
         O(;
         L     #Temp_PV.PV_SetV.WarningUpperLimit;
         L     0.0;
         <=R;
         );
         O(;
         L     #Temp_PV.PV_SetV.Value;
         L     #Temp_PV.PV_SetV.WarningUpperLimit;
         +R;
         L     #Temp_PV.PV_ActV.Value;
         >R;
         );
         JC    gwon;

         L     4;
         T     #Temp_PV.PV_ActV.ValueState;

         JU    end;

   gwon: NOP   0;

   end:  NOP   0;
END_REGION

REGION Network 4: Detect fault levels
   ENDC: O(;
         L     #Temp_PV.PV_ActV.ValueState;
         L     1;
         AW;
         L     0;
         >I;
         );
         AN    #IO_Fault_Alarm_lowerL;
         S     #IO_Fault_Alarm_lowerL;
         S     #IO_New_Fault;

         O(;
         L     #Temp_PV.PV_ActV.ValueState;
         L     2;
         AW;
         L     0;
         >I;
         );
         AN    #IO_Fault_Warn_lowerL;
         S     #IO_Fault_Warn_lowerL;
         S     #IO_New_Fault;

         O(;
         L     #Temp_PV.PV_ActV.ValueState;
         L     4;
         AW;
         L     0;
         >I;
         );
         AN    #IO_Fault_Warn_upperL;
         S     #IO_Fault_Warn_upperL;
         S     #IO_New_Fault;

         O(;
         L     #Temp_PV.PV_ActV.ValueState;
         L     8;
         AW;
         L     0;
         >I;
         );
         AN    #IO_Fault_Alarm_upperL;
         S     #IO_Fault_Alarm_upperL;
         S     #IO_New_Fault;

         O     #IO_Fault_Alarm_lowerL;
         O     #IO_Fault_Alarm_upperL;
         S     #IO_Fault_Level_1;

         O     #IO_Fault_Warn_lowerL;
         O     #IO_Fault_Warn_upperL;
         S     #IO_Fault_Level_3;
END_REGION

REGION Network 5: Write actual value to DB
         CALL  BLKMOV
         ( SRCBLK  := #Temp_PV,
           RET_VAL := #RetVal,
           DSTBLK  := #Anyzeiger_PV
         );
END_REGION
END_FUNCTION

FUNCTION "FC920_PV_Calc_Act_Value" : Void   // FC920, STL
TITLE = Calculates the actual process value of a source
{ S7_Optimized_Access := 'FALSE' }
AUTHOR : HK
VERSION : 0.1
   VAR_INPUT
      IN_Act_Value_read : Bool;   // Read actual value 0 = NO, 1 = YES
      IN_Act_Value_ext : Bool;   // Get actual value from extern
      IN_Ext_Value : Real;   // External value DWord
      IN_Read_Double : Bool;   // Read double word value
      IN_FLT_Needful : Bool;   // Is a seperat fault identification needful?
      IN_FLT_Reset : Bool;
   END_VAR
   VAR_IN_OUT
      IO_Any_ArrayPV : ANY;
      IO_Fault_Sensor : Bool;
      IO_New_Fault : Bool;
      IO_FLT_Level_3 : Bool;
   END_VAR
   VAR_TEMP
      RetVal : Int;
      Anz_BytePV_Act : Int;
      DB_Nr_PV_Act : Int;
      Anyzeiger_Act : ANY;
      Anf_1_PV_Act : Byte;
      Anf_2_PV_Act : Word;
      Temp_PV : "UDT910_ProcessValue";
      Temp_ActV_Pointer : DWord;
      Temp_Fault_Sensor : Bool;
      Temp_CheckSensor : Bool;
   END_VAR
BEGIN

REGION Network 1: Read Array[No_Array] actual value conf. and actual value
         L;  // Pointer auf das Arrays
         LAR1;

         L     W[AR1, P#2.0];  // #Anz_Byte Baugruppe
         T     #Anz_BytePV_Act;

         L     W[AR1, P#4.0];
         T     #DB_Nr_PV_Act;  // DB no prozessvalue actual value

         L     B[AR1, P#7.0];
         T     #Anf_1_PV_Act;

         L     W[AR1, P#8.0];
         T     #Anf_2_PV_Act;  // Start DW prozessvalue actual value [0]

   //
         LAR1;
         L     16#1002;  // Bytes
         T     W[AR1, P#0.0];
         L     #Anz_BytePV_Act;  // Amount of bytes
         T     W[AR1, P#2.0];
         L     #DB_Nr_PV_Act;  // Block no,
         T     W[AR1, P#4.0];
         L     16#84;
         T     LB[AR1, P#6.0];
         L     #Anf_1_PV_Act;
         T     LB[AR1, P#7.0];
         L     #Anf_2_PV_Act;
         T     LW[AR1, P#8.0];

   //
         CALL  BLKMOV
         ( SRCBLK  := #Anyzeiger_Act,
           RET_VAL := #RetVal,
           DSTBLK  := #Temp_PV
         );
   //

   //------- Reset fault -----------------------
         A     #IN_FLT_Reset;
         ON    #IN_FLT_Needful;
         R     #IO_Fault_Sensor;
END_REGION

REGION Network 2: Reset process value
         L     0;
         T     #Temp_PV.PV_ActV.Value;
   //-----
         AN    #IN_Act_Value_read;
         JC    end6;
   //-------------------------------------------
         A     #IN_Act_Value_ext;  // Value is set external
         A     #IN_Act_Value_read;
         JC    extv;
   //-------------------------------------------
         L     #Temp_PV.PV_Conf_ActV.Address;
         L     0;
         ==I;
         JC    end6;
   //-----
END_REGION

REGION Network 3: Calculate actual value

         A     #IN_Act_Value_ext;  // Value is set external
         JC    extv;
   //-------------------------------------------

         L     #Temp_PV.PV_Conf_ActV.Address;
         SLD   3;
         T     #Temp_ActV_Pointer;

         AN    #IN_Read_Double;
         JC    word;
         L     PID[ #Temp_ActV_Pointer];
         T     #Temp_PV.PV_ActV.Value;
         JU    nw02;
   word: L     PIW[ #Temp_ActV_Pointer];
         ITD;
         DTR;
         T     #Temp_PV.PV_ActV.Value;
         JU    nw02;

   extv: L     #IN_Ext_Value;
         T     #Temp_PV.PV_ActV.Value;

   nw02: L     #Temp_PV.PV_Conf_ActV.Multiplier;
         L     0.0;
         ==R;
         JC    nw03;
         L     #Temp_PV.PV_ActV.Value;
         L     #Temp_PV.PV_Conf_ActV.OffsetSignal;
         ITD;
         DTR;
         -R;
         L     #Temp_PV.PV_Conf_ActV.Multiplier;
         /R;
         T     #Temp_PV.PV_ActV.Value;
END_REGION

REGION Network 4: Limit control sensor value if limits <> 0
   nw03: L     #Temp_PV.PV_Conf_ActV.MaxValueSensor;
         L     #Temp_PV.PV_Conf_ActV.MinValueSensor;
         OW;
         L     0;
         <>D;
         =     #Temp_CheckSensor;

         O(;
         L     #Temp_PV.PV_ActV.Value;
         L     #Temp_PV.PV_Conf_ActV.MaxValueSensor;
         >R;
         );
         O(;
         L     #Temp_PV.PV_ActV.Value;
         L     #Temp_PV.PV_Conf_ActV.MinValueSensor;
         <R;
         );
         A     #Temp_CheckSensor;
         =     #Temp_Fault_Sensor;

         AN    #IN_FLT_Needful;
         JC    ResetValue;

         A     #Temp_Fault_Sensor;
         AN    #IO_Fault_Sensor;
         S     #IO_Fault_Sensor;
         S     #IO_New_Fault;

         O     #IO_Fault_Sensor;
         A     #IN_FLT_Needful;
         S     #IO_FLT_Level_3;
         JU    ResetValue;

   NSepFault:NOP   0;
         A     #Temp_Fault_Sensor;
         =     #IO_Fault_Sensor;

   ResetValue:NOP   0;
         AN    #Temp_Fault_Sensor;
         JC    end6;
         L     0.0;
         T     #Temp_PV.PV_ActV.Value;
         JU    end6;
END_REGION

REGION Network 5: Write actual value to DB
   end6: CALL  BLKMOV
         ( SRCBLK  := #Temp_PV,
           RET_VAL := #RetVal,
           DSTBLK  := #Anyzeiger_Act
         );
END_REGION
END_FUNCTION

FUNCTION "CHCKPNCONN" : Void   // FC1001, SCL
{ S7_Optimized_Access := 'FALSE' }
VERSION : 0.1
   VAR_IN_OUT
      GOON : Bool;
      Active : Bool;
      Address : Hw_Io;
      PN_Request : Bool;
      PN_Fault : Bool;
      DONE : Bool;
   END_VAR
   VAR_TEMP
      SLZ_Header : Struct
         LENTHDR : Word;
         N_DR : Word;
      END_STRUCT;
      Dataset : "SZL-IDW#16#xy96_DataSet";
      ReturnValue : Word;
      ReturnValue_1 : Int;
      ReturnHW : Int;
      HW_Kennung : Hw_Io;
      TempAddress : Hw_Io;
      HW_KennungDevice : Hw_SubModule;
      variant_inout : Variant;
   END_VAR
BEGIN
   IF NOT #GOON THEN
       #DONE := false;
   END_IF;

   IF #Active THEN
       IF #GOON AND NOT #DONE THEN

           "PN_Get_DIAG".returnValue := GET_DIAG(MODE := "PN_Get_DIAG".diagMODE, LADDR := #Address,
                                                 CNT_DIAG => "PN_Get_DIAG".CountDiagDetails,
                                                 DIAG := "PN_Get_DIAG".Diag,
                                                 DETAIL :=#variant_inout);

           IF "Flag_Req_read_IO_Busy" = 0 THEN
               // Bearbeitung beendet
               #DONE := true;
               // Fehler wurde festgestellt
               IF ("PN_Get_DIAG".Diag.OwnState > 0)

               THEN
                   #PN_Fault := true;
                   #PN_Request := false;
               END_IF;
               // Fehler wurde behoben
               IF #PN_Fault AND ("PN_Get_DIAG".Diag.OwnState = 0)

               THEN
                   #PN_Request := true;//#PN_Fault;
                   #PN_Fault := false;
               END_IF;
           END_IF;
       END_IF;
   ELSE
       #DONE := #GOON;
   END_IF;
   // Zusätzlichen Ausgang schreiben
   // 
   #GOON := #DONE;



   // Unten ist der alte Code
   // IF #GoOn THEN
   //     #ReturnValue := INT_TO_WORD(RDSYSST(REQ := true, //"Flag_01_000_Hertz" ,
   //                                                                     SZL_ID := 16#0696,
   //                                                                     INDEX := DINT_TO_WORD(#Address),
   //                                                                     BUSY => "Flag_Req_read_DP1_Busy",
   //                                                                     SZL_HEADER => #SLZ_Header,
   //                                                                     DR => "PN_CON".Dataset));

   //     IF #ReturnValue <> 0 THEN
   //         IF (NOT "PN_CON".Dataset.IOStat.BaugruppeVorhanden) OR "PN_CON".Dataset.IOStat.BaugruppeDeaktiviert OR "PN_CON".Dataset.IOStat.BaugruppeNichtVerfuegbar THEN

   //             #PN_Fault := true;
   //             #PN_Request := false;
   //         END_IF;

   //         IF #PN_Fault AND "PN_CON".Dataset.IOStat.BaugruppeVorhanden AND NOT "PN_CON".Dataset.IOStat.BaugruppeDeaktiviert AND NOT "PN_CON".Dataset.IOStat.BaugruppeNichtVerfuegbar THEN
   //             #PN_Request := true;
   //             #PN_Fault := false;
   //         END_IF;
   //     END_IF;
   //     IF WORD_TO_INT(#ReturnValue) > 16#8000 THEN
   //             #PN_Fault := true;
   //     END_IF;
   // END_IF;
END_FUNCTION

FUNCTION "PNC_AI" : Void   // FC1002, SCL
{ S7_Optimized_Access := 'FALSE' }
VERSION : 0.1
   VAR_INPUT
      RequestAll : Bool;
      AcknowledgeFaults : Bool;
   END_VAR
   VAR_IN_OUT
      GOON : Bool;
   END_VAR
   VAR_TEMP
      t : Struct
         DONE : Bool;
         BUSY : Bool;
         ERROR : Bool;
         STATUS : DWord;
      END_STRUCT;
      MODULE : Int;
      ADDRESS : Word;
      MinIndex : Int;
      MaxIndex : Int;
      SLZ_Header : Struct
         LENTHDR : Word;
         N_DR : Word;
      END_STRUCT;
      Dataset : "SZL-IDW#16#xy96_DataSet";
      TempHWID : Hw_Io;
      ReturnValue : Int;
   END_VAR
   VAR CONSTANT
      IDM_Analogin_Default_Skalierung_Index : Int := 2;
      IDM_Analogin_Default_Skalierung_Length : Int := 4;
      IDM_Analogin_Default_Filterung_Index : Int := 3;
      IDM_Analogin_Default_Filterung_Length : Int := 2;
      IDM_Analogin_Default_Grenzen_Index : Int := 4;
      IDM_Analogin_Default_Grenzen_Length : Int := 12;
      IDM_Analogin_Default_8_X14_0_Index : Int := 1;
      IDM_Analogin_Default_8_X14_0_Length : Int := 64;
      IDM_Analogin_Temperature_Index : Int := 2;
      IDM_Analogin_Temperature_Length : Int := 5;
      IDM_Analogin_Temperature_8_Index : Int := 1;
      IDM_Analogin_Temperature_8_Length : Int := 48;
   END_VAR
BEGIN
   // Setze Grenzen für das Durchlaufen der Schleife
   // 
   #MinIndex := 1;
   #MaxIndex := 16;

   // Überwachung des maximalen Index
   // 
   IF #AcknowledgeFaults THEN
       "PN_AI".IndexError := false;
   END_IF;
   IF #MaxIndex > 16 THEN
       #MaxIndex := 16;
       "PN_AI".IndexError := true;
   END_IF;

   // -----------------------------
   // Schnittstelle für Visualisierung (Modulauswahl)
   // -----------------------------
   IF "PN_AI".SetIndex > #MaxIndex THEN
       "PN_AI".SetIndex := #MinIndex;
   ELSIF "PN_AI".SetIndex < #MinIndex THEN
       "PN_AI".SetIndex := #MaxIndex;
   END_IF;

   IF ("PN_AI".SetIndex <> "PN_AI".ActIndex) OR "PN_AI".Send THEN
       "PN_AI".Module["PN_AI".ActIndex] := "PN_AI".Module[0];
       "PN_AI".Module[0] := "PN_AI".Module["PN_AI".SetIndex];
       "PN_AI".ActIndex := "PN_AI".SetIndex;
       "PN_AI".Send := false;
   END_IF;

   // -----------------------------
   // Verschicken der Telegramme
   // -----------------------------
   FOR #MODULE := #MinIndex TO #MaxIndex DO
       IF #RequestAll = true THEN
           "PN_AI".Module[#MODULE].AI8.X14_0.Request := "PN_AI".Module[#MODULE].AI8.Active;
           "PN_AI".Module[#MODULE].AIResistive_8.TemperatureInput.Request := "PN_AI".Module[#MODULE].AIResistive_8.Active;
       END_IF;

       // Wenn ein Modul nicht aktiviert ist, dann soll auch der Request zurückgesetzt werden.
       IF (NOT "PN_AI".Module[#MODULE].AI8.Active) OR
           ("PN_AI".Module[#MODULE].AI8.Address = 0)
       THEN
           "PN_AI".Module[#MODULE].AI8.X14_0.Request := false;
       END_IF;
       IF (NOT "PN_AI".Module[#MODULE].AIResistive_8.Active) OR
           ("PN_AI".Module[#MODULE].AIResistive_8.Address = 0)
       THEN
           "PN_AI".Module[#MODULE].AIResistive_8.TemperatureInput.Request := false;
       END_IF;

       // Paremetrierung der Analogen Eingänge
       // 
       #ADDRESS := INT_TO_WORD("PN_AI".Module[#MODULE].AI8.Address);
       #ReturnValue := LOG2MOD(IOID := B#16#54, ADDR := #ADDRESS, HWID => #TempHWID);
       // Kommunikationsüberwachung
       // Nach einem Verbindungsabbruch werden die Telegramme automatisch verschickt.
       "CHCKPNCONN"(GOON := #GOON,
                    Active := "PN_AI".Module[#MODULE].AI8.Active,
                    Address := #TempHWID,
                    PN_Request := "PN_AI".Module[#MODULE].AI8.X14_0.Request,
                    PN_Fault := "PN_AI".Module[#MODULE].AI8.ChckConnFault,
                    DONE := "PN_AI".Module[#MODULE].AI8.ChckConnDone);

       "WRREC_FC"(GOON := #GOON,
                  REQ := "PN_AI".Module[#MODULE].AI8.X14_0.Request,
                  ADDRESS := #TempHWID,
                  INDEX := #IDM_Analogin_Default_8_X14_0_Index,
                  LENGTH := #IDM_Analogin_Default_8_X14_0_Length,
                  WRREC_DONE => #t.DONE,
                  WRREC_BUSY => #t.BUSY,
                  WRREC_ERROR => #t.ERROR,
                  WRREC_STATUS => #t.STATUS,
                  ACTIVE := "PN_AI".Module[#MODULE].AI8.Active,
                  RECORD := "PN_AI".Module[#MODULE].AI8.X14_0.Data,
                  DONE := "PN_AI".Module[#MODULE].AI8.X14_0.Transmitting);

       // Parametrierung der Analogen Temperatur Eingänge
       #ADDRESS := INT_TO_WORD("PN_AI".Module[#MODULE].AIResistive_8.Address);
       #ReturnValue := LOG2MOD(IOID := B#16#54, ADDR := #ADDRESS, HWID => #TempHWID);
       // Kommunikationsüberwachung
       // Nach einem Verbindungsabbruch werden die Telegramme automatisch verschickt.
       "CHCKPNCONN"(GOON := #GOON,
                    Active := "PN_AI".Module[#MODULE].AIResistive_8.Active,
                    Address := #TempHWID,
                    PN_Request := "PN_AI".Module[#MODULE].AIResistive_8.TemperatureInput.Request,
                    PN_Fault := "PN_AI".Module[#MODULE].AIResistive_8.ChckConnFault,
                    DONE := "PN_AI".Module[#MODULE].AIResistive_8.ChckConnDone);

       "WRREC_FC"(GOON := #GOON,
                  REQ := "PN_AI".Module[#MODULE].AIResistive_8.TemperatureInput.Request,
                  ADDRESS := #TempHWID,
                  INDEX := #IDM_Analogin_Temperature_8_Index,
                  LENGTH := #IDM_Analogin_Temperature_8_Length,
                  WRREC_DONE => #t.DONE,
                  WRREC_BUSY => #t.BUSY,
                  WRREC_ERROR => #t.ERROR,
                  WRREC_STATUS => #t.STATUS,
                  ACTIVE := "PN_AI".Module[#MODULE].AIResistive_8.Active,
                  RECORD := "PN_AI".Module[#MODULE].AIResistive_8.TemperatureInput.Data,
                  DONE := "PN_AI".Module[#MODULE].AIResistive_8.TemperatureInput.Transmitting);
   END_FOR;
END_FUNCTION

FUNCTION "PNC_Flow" : Void   // FC1003, SCL
{ S7_Optimized_Access := 'FALSE' }
VERSION : 0.1
   VAR_INPUT
      RequestAll : Bool;
      AcknowledgeFaults : Bool;
   END_VAR
   VAR_IN_OUT
      GOON : Bool;
   END_VAR
   VAR_TEMP
      t : Struct
         DONE : Bool;
         BUSY : Bool;
         ERROR : Bool;
         STATUS : DWord;
      END_STRUCT;
      ADDRESS : Word;
      "COUNTER" : Int;
      MinIndex : Int;
      MaxIndex : Int;
      dummy : Real;
      Request : Bool;
      TempHWID : Hw_Io;
      ReturnValue : Int;
      ExternSetting : Bool;
      TempGOON : Bool;
   END_VAR
   VAR CONSTANT
      IDM_Analogout_Flow_Controller_HardwareResourcen_Index : Int := 1;
      IDM_Analogout_Flow_Controller_HardwareResourcen_Length : Int := 10;
      IDM_Analogout_Flow_Controller_GeneralParameters_Index : Int := 2;
      IDM_Analogout_Flow_Controller_GeneralParameters_Length : Int := 16;
      IDM_Analogout_Flow_Controller_Grenzen_Index : Int := 3;
      IDM_Analogout_Flow_Controller_Grenzen_Length : Int := 16;
      IDM_Analogout_Flow_Controller_Skalierung_Index : Int := 4;
      IDM_Analogout_Flow_Controller_Skalierung_Length : Int := 12;
      IDM_FlowSpeed_Skalierung_Index : Int := 2;
      IDM_FlowSpeed_Skalierung_Length : Int := 6;
   END_VAR
BEGIN

   // -----------------------------
   // Telegrammübermittlung
   // -----------------------------
   #MinIndex := 1;
   #MaxIndex := 4;
   #ExternSetting := FALSE;

   FOR #COUNTER := #MinIndex TO #MaxIndex DO

       IF "DB900_ConfCalibFlow".Flow[#COUNTER].Density <> "DB702_Tank_Value".Tank["DB753_MeteringPump".Pump[#COUNTER].TankNo].Density THEN
           "DB900_ConfCalibFlow".Flow[#COUNTER].Density := "DB702_Tank_Value".Tank["DB753_MeteringPump".Pump[#COUNTER].TankNo].Density;
           "PN_FlowRate".Component[#COUNTER].FlowC_F.GeneralParameters.Request := true;
           #ExternSetting := TRUE;
       END_IF;
       IF "DB900_ConfCalibFlow".Flow[#COUNTER].Factor <> "DB753_MeteringPump".Pump[#COUNTER].FlowFactor THEN
           "DB900_ConfCalibFlow".Flow[#COUNTER].Factor := "DB753_MeteringPump".Pump[#COUNTER].FlowFactor;
           "PN_FlowRate".Component[#COUNTER].FlowC_F.GeneralParameters.Request := true;
           #ExternSetting := TRUE;
       END_IF;
       IF "DB900_ConfCalibFlow".Flow[#COUNTER].Pulse_per_liter <> "DB753_MeteringPump".Pump[#COUNTER].Pulse_per_liter THEN
           "DB900_ConfCalibFlow".Flow[#COUNTER].Pulse_per_liter := "DB753_MeteringPump".Pump[#COUNTER].Pulse_per_liter;
           "PN_FlowRate".Component[#COUNTER].FlowC_F.GeneralParameters.Request := true;
           #ExternSetting := TRUE;
       END_IF;
       IF "DB900_ConfCalibFlow".Flow[#COUNTER].MaxFlow <> "DB613_Komponent_State".FlowPumpMax[#COUNTER] THEN
           "DB900_ConfCalibFlow".Flow[#COUNTER].MaxFlow := "DB613_Komponent_State".FlowPumpMax[#COUNTER];
           "PN_FlowRate".Component[#COUNTER].FlowC_F.GeneralParameters.Data.MaxDurchfluss := "DB900_ConfCalibFlow".Flow[#COUNTER].MaxFlow;
           "PN_FlowRate".Component[#COUNTER].FlowC_F.GeneralParameters.Request := true;
           #ExternSetting := TRUE;
       END_IF;

       "PN_FlowRate".Component[#COUNTER].FlowC_F.GeneralParameters.Data.Kalibrierfaktor :=
       INT_TO_REAL("DB702_Tank_Value".Tank["DB753_MeteringPump".Pump[#COUNTER].TankNo].Density) /
       "DB753_MeteringPump".Pump[#COUNTER].Pulse_per_liter *
       "DB753_MeteringPump".Pump[#COUNTER].FlowFactor;

       IF #ExternSetting = TRUE AND "PN_FlowRate".SetIndex = #COUNTER THEN
           "PN_FlowRate".Component[0] := "PN_FlowRate".Component["PN_FlowRate".SetIndex];
       END_IF;

   END_FOR;

   IF #AcknowledgeFaults THEN
       "PN_FlowRate".IndexError := false;
   END_IF;
   IF #MaxIndex > 16 THEN
       #MaxIndex := 16;
       "PN_FlowRate".IndexError := true;
   END_IF;

   // Calculate the Parameter bits to the konfiguration Byte
   "PN_FlowRate".Component[0].FlowC_F.Hardware.Data.Konfig1 :=
   SHL(IN := "PN_FlowRate".Component[0].FlowC_F.Visualisierung.BetriebsartAnalogausgang, N := 0) OR
   SHL(IN := "PN_FlowRate".Component[0].FlowC_F.Visualisierung.BipolarerAusgang, N := 3) OR
   SHL(IN := "PN_FlowRate".Component[0].FlowC_F.Visualisierung.Polarität, N := 4) OR
   SHL(IN := "PN_FlowRate".Component[0].FlowC_F.Visualisierung.BetriebsartAnalogeingang, N := 5);

   "PN_FlowRate".Component[0].FlowC_F.Hardware.Data.Konfig2 :=
   SHL(IN := "PN_FlowRate".Component[0].FlowC_F.Visualisierung.BetriebsartQuadraturdekoder, N := 0) OR
   SHL(IN := "PN_FlowRate".Component[0].FlowC_F.Visualisierung.QuelleIstdruck, N := 3);

   // -----------------------------
   // Schnittstelle für Visualisierung
   // -----------------------------
   IF "PN_FlowRate".SetIndex > #MaxIndex THEN
       "PN_FlowRate".SetIndex := #MinIndex;
   ELSIF "PN_FlowRate".SetIndex < #MinIndex THEN
       "PN_FlowRate".SetIndex := #MaxIndex;
   END_IF;

   IF ("PN_FlowRate".SetIndex <> "PN_FlowRate".ActIndex) OR "PN_FlowRate".Send THEN
       "PN_FlowRate".Component["PN_FlowRate".ActIndex] := "PN_FlowRate".Component[0];
       "PN_FlowRate".Component[0] := "PN_FlowRate".Component["PN_FlowRate".SetIndex];
       "PN_FlowRate".ActIndex := "PN_FlowRate".SetIndex;
       "PN_FlowRate".Send := false;
   END_IF;

   // -----------------------------
   // Prüfe die Anforderungen (Request)
   // -----------------------------
   FOR #COUNTER := #MinIndex TO #MaxIndex DO

       // Calculate the Parameter bits to the konfiguration Byte
       "PN_FlowRate".Component[#COUNTER].FlowC_F.Hardware.Data.Konfig1 :=
       SHL(IN := "PN_FlowRate".Component[#COUNTER].FlowC_F.Visualisierung.BetriebsartAnalogausgang, N := 0) OR
       SHL(IN := "PN_FlowRate".Component[#COUNTER].FlowC_F.Visualisierung.BipolarerAusgang, N := 3) OR
       SHL(IN := "PN_FlowRate".Component[#COUNTER].FlowC_F.Visualisierung.Polarität, N := 4) OR
       SHL(IN := "PN_FlowRate".Component[#COUNTER].FlowC_F.Visualisierung.BetriebsartAnalogeingang, N := 5);

       "PN_FlowRate".Component[#COUNTER].FlowC_F.Hardware.Data.Konfig2 :=
       SHL(IN := "PN_FlowRate".Component[#COUNTER].FlowC_F.Visualisierung.BetriebsartQuadraturdekoder, N := 0) OR
       SHL(IN := "PN_FlowRate".Component[#COUNTER].FlowC_F.Visualisierung.QuelleIstdruck, N := 3);

       IF #RequestAll = TRUE THEN
           //        "PN_FlowRate".Component[#COUNTER].FlowC_F.Hardware.Request := "PN_FlowRate".Component[#COUNTER].FlowC_F.Active;
           "PN_FlowRate".Component[#COUNTER].FlowC_F.GeneralParameters.Request := "PN_FlowRate".Component[#COUNTER].FlowC_F.Active;
           "PN_FlowRate".Component[#COUNTER].FlowC_F.Grenzen.Request := "PN_FlowRate".Component[#COUNTER].FlowC_F.Active;
           "PN_FlowRate".Component[#COUNTER].FlowC_F.SkalierungAI.Request := "PN_FlowRate".Component[#COUNTER].FlowC_F.Active;
           //        "PN_FlowRate".Component[#COUNTER].Flow_F.Skalierung.Request := true;
       END_IF;
       // Wenn ein Modul nicht aktiviert ist, dann soll auch der Request zurückgesetzt werden.
       IF (NOT "PN_FlowRate".Component[#COUNTER].FlowC_F.Active) OR
           ("PN_FlowRate".Component[#COUNTER].FlowC_F.Address = 0)
       THEN
           "PN_FlowRate".Component[#COUNTER].FlowC_F.Hardware.Request := false;
           "PN_FlowRate".Component[#COUNTER].FlowC_F.GeneralParameters.Request := false;
           "PN_FlowRate".Component[#COUNTER].FlowC_F.Grenzen.Request := false;
           "PN_FlowRate".Component[#COUNTER].FlowC_F.SkalierungAI.Request := false;
       END_IF;
       // ======================================================================================
       // Durchflussregler 
       // ======================================================================================
       "PN_FlowRate".Component[1].FlowC_F.Address := 1000;
       "PN_FlowRate".Component[2].FlowC_F.Address := 1100;

       #ADDRESS := INT_TO_WORD("PN_FlowRate".Component[#COUNTER].FlowC_F.Address);
       #ReturnValue := LOG2MOD(IOID := B#16#54, ADDR := #ADDRESS, HWID => #TempHWID);
       // Kommunikationsüberwachung
       // Nach einem Verbindungsabbruch werden die Telegramme automatisch verschickt.
       #Request := false;
       "CHCKPNCONN"(GOON := #GOON,
                    Active := "PN_FlowRate".Component[#COUNTER].FlowC_F.Active,
                    Address := #TempHWID,
                    PN_Request := #Request,
                    PN_Fault := "PN_FlowRate".Component[#COUNTER].FlowC_F.ChckConnFault,
                    DONE := "PN_FlowRate".Component[#COUNTER].FlowC_F.ChckConnDone);

       IF #Request AND NOT "PN_FlowRate".Component[#COUNTER].FlowC_F.ChckConnFault THEN
           //        "PN_FlowRate".Component[#COUNTER].FlowC_F.Hardware.Request := "PN_FlowRate".Component[#COUNTER].FlowC_F.Active;
           "PN_FlowRate".Component[#COUNTER].FlowC_F.GeneralParameters.Request := "PN_FlowRate".Component[#COUNTER].FlowC_F.Active;
           "PN_FlowRate".Component[#COUNTER].FlowC_F.Grenzen.Request := "PN_FlowRate".Component[#COUNTER].FlowC_F.Active;
           "PN_FlowRate".Component[#COUNTER].FlowC_F.SkalierungAI.Request := "PN_FlowRate".Component[#COUNTER].FlowC_F.Active;
       END_IF;

   //    #TempGOON:= #GOON AND NOT ("PN_FlowRate".Component[#COUNTER].FlowC_F.Grenzen.Busy OR "PN_FlowRate".Component[#COUNTER].FlowC_F.SkalierungAI.Busy)

       "WRREC_FC"(GOON := #GOON,
                  REQ := "PN_FlowRate".Component[#COUNTER].FlowC_F.GeneralParameters.Request,
                  ADDRESS := #TempHWID,
                  INDEX := #IDM_Analogout_Flow_Controller_GeneralParameters_Index,
                  LENGTH := #IDM_Analogout_Flow_Controller_GeneralParameters_Length,
                  WRREC_DONE => "PN_FlowRate".Component[#COUNTER].FlowC_F.GeneralParameters.Done,
                  WRREC_BUSY => "PN_FlowRate".Component[#COUNTER].FlowC_F.GeneralParameters.Busy,
                  WRREC_ERROR => #t.ERROR,
                  WRREC_STATUS => #t.STATUS,
                  ACTIVE := "PN_FlowRate".Component[#COUNTER].FlowC_F.Active,
                  RECORD := "PN_FlowRate".Component[#COUNTER].FlowC_F.GeneralParameters.Data,
                  DONE := "PN_FlowRate".Component[#COUNTER].FlowC_F.GeneralParameters.Transmitting);

       "WRREC_FC"(GOON := #GOON,
                  REQ := "PN_FlowRate".Component[#COUNTER].FlowC_F.Grenzen.Request,
                  ADDRESS := #TempHWID,
                  INDEX := #IDM_Analogout_Flow_Controller_Grenzen_Index,
                  LENGTH := #IDM_Analogout_Flow_Controller_Grenzen_Length,
                  WRREC_DONE => "PN_FlowRate".Component[#COUNTER].FlowC_F.Grenzen.Done,
                  WRREC_BUSY => "PN_FlowRate".Component[#COUNTER].FlowC_F.Grenzen.Busy,
                  WRREC_ERROR => #t.ERROR,
                  WRREC_STATUS => #t.STATUS,
                  ACTIVE := "PN_FlowRate".Component[#COUNTER].FlowC_F.Active,
                  RECORD := "PN_FlowRate".Component[#COUNTER].FlowC_F.Grenzen.Data,
                  DONE := "PN_FlowRate".Component[#COUNTER].FlowC_F.Grenzen.Tranmitting);

       "WRREC_FC"(GOON := #GOON,
                  REQ := "PN_FlowRate".Component[#COUNTER].FlowC_F.SkalierungAI.Request,
                  ACTIVE := "PN_FlowRate".Component[#COUNTER].FlowC_F.Active,
                  ADDRESS := #TempHWID,
                  INDEX := #IDM_Analogout_Flow_Controller_Skalierung_Index,
                  LENGTH := #IDM_Analogout_Flow_Controller_Skalierung_Length,
                  WRREC_DONE => "PN_FlowRate".Component[#COUNTER].FlowC_F.SkalierungAI.Done,
                  WRREC_BUSY => "PN_FlowRate".Component[#COUNTER].FlowC_F.SkalierungAI.Busy,
                  WRREC_ERROR => #t.ERROR,
                  WRREC_STATUS => #t.STATUS,
                  RECORD := "PN_FlowRate".Component[#COUNTER].FlowC_F.SkalierungAI.Data,
                  DONE := "PN_FlowRate".Component[#COUNTER].FlowC_F.SkalierungAI.Transmitting);

       // ======================================================================================
       // Durchfluss OHNE Regler
       // ======================================================================================
       #ADDRESS := INT_TO_WORD("PN_FlowRate".Component[#COUNTER].FlowC_F.Address);
       #ReturnValue := LOG2MOD(IOID := B#16#54, ADDR := #ADDRESS, HWID => #TempHWID);
       // Kommunikationsüberwachung
       // Nach einem Verbindungsabbruch werden die Telegramme automatisch verschickt.
       #Request := false;
       "CHCKPNCONN"(GOON := #GOON,
                    Active := "PN_FlowRate".Component[#COUNTER].Flow_F.Active,
                    Address := #TempHWID,
                    PN_Request := #Request,
                    PN_Fault := "PN_FlowRate".Component[#COUNTER].Flow_F.ChckConnFault,
                    DONE := "PN_FlowRate".Component[#COUNTER].Flow_F.ChckConnDone);

       IF #Request AND NOT "PN_FlowRate".Component[#COUNTER].Flow_F.ChckConnFault THEN
           "PN_FlowRate".Component[#COUNTER].Flow_F.Skalierung.Request := "PN_FlowRate".Component[#COUNTER].Flow_F.Active;
       END_IF;
       // "WRREC_FC"(REQ := "PN_FlowRate".Component[#COUNTER].Flow_F.Skalierung.Request,
       //            TRANSMITTING := "PN_FlowRate".Component[#COUNTER].Flow_F.Skalierung.Transmitting,
       //             ADDRESS := #TempHWID,
       //             INDEX := #IDM_FlowSpeed_Skalierung_Index,s
       //             LENGTH := #IDM_FlowSpeed_Skalierung_Length,
       //             DONE => #t.DONE,
       //             BUSY => #t.BUSY,
       //             ERROR => #t.ERROR,
       //             STATUS => #t.STATUS,
       //             ACTIVE:=#COMPONENT[#COUNTER].FLOW.ACTIVE,
       //             RECORD := "PN_FlowRate".Component[#COUNTER].Flow_F.Skalierung.Data);
   END_FOR;
END_FUNCTION

FUNCTION "PNC_Mixinghead" : Void   // FC1004, SCL
{ S7_Optimized_Access := 'FALSE' }
VERSION : 0.1
   VAR_INPUT
      RequestAll : Bool;
      AcknowledgeFaults : Bool;
   END_VAR
   VAR_IN_OUT
      GOON : Bool;
   END_VAR
   VAR_TEMP
      t : Struct
         DONE : Bool;
         BUSY : Bool;
         ERROR : Bool;
         STATUS : DWord;
      END_STRUCT;
      MH : Int;   // Mischkopfzähler
      DB : Int;   // Düse/Bypass-Zähler
      Address : Word;
      MinIndex : Int;
      MaxIndex : Int;
      Request : Bool;
      TempHWID : Hw_Io;
      ReturnValue : Int;
      Fault : Bool;
   END_VAR
   VAR CONSTANT
      IDM_Mixinghead_Digital_GeneralParameters_Index : Int := 1;
      IDM_Mixinghead_Digital_GeneralParameters_Length : Int := 4;
      IDM_Mixinghead_Digital_Zeiten_Index : Int := 2;
      IDM_Mixinghead_Digital_Zeiten_Length : Int := 12;
      IDM_Mixinghead_Digital_Zeiten_2_Index : Int := 6;
      IDM_Mixinghead_Digital_Zeiten_2_Length : Int := 4;
      IDM_Mixinghead_Analog_Resourcen_Index : Int := 1;
      IDM_Mixinghead_Analog_Resourcen_Length : Int := 8;
      IDM_Mixinghead_Analog_Zeiten_Index : Int := 2;
      IDM_Mixinghead_Analog_Zeiten_Length : Int := 6;
      IDM_Mixinghead_Analog_Skalierung_Index : Int := 3;
      IDM_Mixinghead_Analog_Skalierung_Length : Int := 4;
      IDM_Mixinghead_Analog_StufenAktivierung_Index : Int := 4;
      IDM_Mixinghead_Analog_StufenAktivierung_Length : Int := 20;
      IDM_Mixinghead_Analog_StufenRückkehr_Index : Int := 5;
      IDM_Mixinghead_Analog_StufenRückkehr_Length : Int := 20;
      IDM_CleaningPiston_Digital_GeneralParameters_Index : Int := 1;
      IDM_CleaningPiston_Digital_GeneralParameters_Length : Int := 3;
      IDM_CleaningPiston_Digital_Zeiten_Index : Int := 2;
      IDM_CleaningPiston_Digital_Zeiten_Length : Int := 20;
      IDM_CleaningPiston_Analog_GeneralParameters_Index : Int := 1;
      IDM_CleaningPiston_Analog_GeneralParameters_Length : Int := 6;
      IDM_CleaningPiston_Analog_Zeiten_Index : Int := 2;
      IDM_CleaningPiston_Analog_Zeiten_Length : Int := 14;
      IDM_CleaningPiston_Analog_Skalierung_Index : Int := 3;
      IDM_CleaningPiston_Analog_Skalierung_Length : Int := 4;
      IDM_CleaningPiston_Analog_StufenAktivierung_Index : Int := 4;
      IDM_CleaningPiston_Analog_StufenAktivierung_Length : Int := 20;
      IDM_CleaningPiston_Analog_StufenRückkehr_Index : Int := 5;
      IDM_CleaningPiston_Analog_StufenRückkehr_Length : Int := 20;
      IDM_CleaningPiston_Analog_Loop_GeneralParameters_Index : Int := 1;
      IDM_CleaningPiston_Analog_Loop_GeneralParameters_Length : Int := 5;
      IDM_CleaningPiston_Analog_Loop_Zeiten_Index : Int := 2;
      IDM_CleaningPiston_Analog_Loop_Zeiten_Length : Int := 14;
      IDM_CleaningPiston_Analog_Loop_Regelparameter_Index : Int := 4;
      IDM_CleaningPiston_Analog_Loop_Regelparameter_Length : Int := 12;
      IDM_Mixinghead_NozzleBypass_Kanal_Index : Int := 1;
      IDM_Mixinghead_NozzleBypass_Kanal_Length : Int := 3;
      IDM_Mixinghead_NozzleBypass_Zeiten_Index : Int := 2;
      IDM_Mixinghead_NozzleBypass_Zeiten_Length : Int := 8;
   END_VAR
BEGIN
   #MinIndex := 1;
   #MaxIndex := 2;

   IF #AcknowledgeFaults THEN
       "PN_Mixinghead".IndexError := false;
   END_IF;
   IF #MaxIndex > 16 THEN
       #MaxIndex := 16;
       "PN_Mixinghead".IndexError := true;
   END_IF;
   // -----------------------------
   // Schnittstelle für Visualisierung
   // -----------------------------
   IF "PN_Mixinghead".SetIndex > #MaxIndex THEN
       "PN_Mixinghead".SetIndex := #MinIndex;
   ELSIF "PN_Mixinghead".SetIndex < #MinIndex THEN
       "PN_Mixinghead".SetIndex := #MaxIndex;
   END_IF;

   IF ("PN_Mixinghead".SetIndex <> "PN_Mixinghead".ActIndex) OR "PN_Mixinghead".Send THEN
       "PN_Mixinghead".Mixinghead["PN_Mixinghead".ActIndex] := "PN_Mixinghead".Mixinghead[0];
       "PN_Mixinghead".Mixinghead[0] := "PN_Mixinghead".Mixinghead["PN_Mixinghead".SetIndex];
       "PN_Mixinghead".ActIndex := "PN_Mixinghead".SetIndex;
       "PN_Mixinghead".Send := false;
   END_IF;

   // -----------------------------
   // Prüfe die Anforderungen (Request)
   // -----------------------------
   FOR #MH := #MinIndex TO #MaxIndex DO
       IF #RequestAll = True THEN
           "PN_Mixinghead".Mixinghead[#MH].Analog.Resourcen.Request := "PN_Mixinghead".Mixinghead[#MH].Analog.Active;
           "PN_Mixinghead".Mixinghead[#MH].Analog.Zeiten.Request := "PN_Mixinghead".Mixinghead[#MH].Analog.Active;
           "PN_Mixinghead".Mixinghead[#MH].Analog.Skalierung.Request := "PN_Mixinghead".Mixinghead[#MH].Analog.Active;
           "PN_Mixinghead".Mixinghead[#MH].Analog.StufenAktivierung.Request := "PN_Mixinghead".Mixinghead[#MH].Analog.Active;
           "PN_Mixinghead".Mixinghead[#MH].Analog.StufenRückkehr.Request := "PN_Mixinghead".Mixinghead[#MH].Analog.Active;

           "PN_Mixinghead".Mixinghead[#MH].Digital.GeneralParameters.Request := "PN_Mixinghead".Mixinghead[#MH].Digital.Active;
           "PN_Mixinghead".Mixinghead[#MH].Digital.Zeiten.Request := "PN_Mixinghead".Mixinghead[#MH].Digital.Active;

           "PN_Mixinghead".Mixinghead[#MH].ReinigungskolbenDigital.GeneralParameters.Request := "PN_Mixinghead".Mixinghead[#MH].ReinigungskolbenDigital.Active;
           "PN_Mixinghead".Mixinghead[#MH].ReinigungskolbenDigital.Zeiten.Request := "PN_Mixinghead".Mixinghead[#MH].ReinigungskolbenDigital.Active;

           "PN_Mixinghead".Mixinghead[#MH].ReinigungskolbenGeregelt.GeneralParameters.Request := "PN_Mixinghead".Mixinghead[#MH].ReinigungskolbenGeregelt.Active;
           "PN_Mixinghead".Mixinghead[#MH].ReinigungskolbenGeregelt.Zeiten.Request := "PN_Mixinghead".Mixinghead[#MH].ReinigungskolbenGeregelt.Active;
           "PN_Mixinghead".Mixinghead[#MH].ReinigungskolbenGeregelt.Skalierung.Request := "PN_Mixinghead".Mixinghead[#MH].ReinigungskolbenGeregelt.Active;
           "PN_Mixinghead".Mixinghead[#MH].ReinigungskolbenGeregelt.Regelparameter.Request := "PN_Mixinghead".Mixinghead[#MH].ReinigungskolbenGeregelt.Active;

           "PN_Mixinghead".Mixinghead[#MH].ReinigungskolbenGesteuert.GeneralParameters.Request := "PN_Mixinghead".Mixinghead[#MH].ReinigungskolbenGesteuert.Active;
           "PN_Mixinghead".Mixinghead[#MH].ReinigungskolbenGesteuert.Zeiten.Request := "PN_Mixinghead".Mixinghead[#MH].ReinigungskolbenGesteuert.Active;
           "PN_Mixinghead".Mixinghead[#MH].ReinigungskolbenGesteuert.Skalierung.Request := "PN_Mixinghead".Mixinghead[#MH].ReinigungskolbenGesteuert.Active;
           "PN_Mixinghead".Mixinghead[#MH].ReinigungskolbenGesteuert.StufenAktivierung.Request := "PN_Mixinghead".Mixinghead[#MH].ReinigungskolbenGesteuert.Active;
           "PN_Mixinghead".Mixinghead[#MH].ReinigungskolbenGesteuert.StufenRückkehr.Request := "PN_Mixinghead".Mixinghead[#MH].ReinigungskolbenGesteuert.Active;
           FOR #DB := 1 TO 8 DO
               "PN_Mixinghead".Mixinghead[#MH].DüseBypass[#DB].Zeiten.Request := "PN_Mixinghead".Mixinghead[#MH].DüseBypass[#DB].Active;
           END_FOR;
       END_IF;

       // Wenn ein Modul nicht aktiviert ist, dann soll auch der Request zurückgesetzt werden.
       IF NOT "PN_Mixinghead".Mixinghead[#MH].Analog.Active OR
           "PN_Mixinghead".Mixinghead[#MH].Analog.Address = 0
       THEN
           "PN_Mixinghead".Mixinghead[#MH].Analog.Resourcen.Request := false;
           "PN_Mixinghead".Mixinghead[#MH].Analog.Zeiten.Request := false;
           "PN_Mixinghead".Mixinghead[#MH].Analog.Skalierung.Request := false;
           "PN_Mixinghead".Mixinghead[#MH].Analog.StufenAktivierung.Request := false;
           "PN_Mixinghead".Mixinghead[#MH].Analog.StufenRückkehr.Request := false;
       END_IF;
       IF NOT "PN_Mixinghead".Mixinghead[#MH].Digital.Active OR
           "PN_Mixinghead".Mixinghead[#MH].Digital.Address = 0
       THEN
           "PN_Mixinghead".Mixinghead[#MH].Digital.GeneralParameters.Request := false;
           "PN_Mixinghead".Mixinghead[#MH].Digital.Zeiten.Request := false;
       END_IF;
       IF NOT "PN_Mixinghead".Mixinghead[#MH].ReinigungskolbenDigital.Active OR
           "PN_Mixinghead".Mixinghead[#MH].ReinigungskolbenDigital.Address = 0
       THEN
           "PN_Mixinghead".Mixinghead[#MH].ReinigungskolbenDigital.GeneralParameters.Request := false;
           "PN_Mixinghead".Mixinghead[#MH].ReinigungskolbenDigital.Zeiten.Request := false;
       END_IF;
       IF NOT "PN_Mixinghead".Mixinghead[#MH].ReinigungskolbenGeregelt.Active OR
           "PN_Mixinghead".Mixinghead[#MH].ReinigungskolbenGeregelt.Address = 0
       THEN
           "PN_Mixinghead".Mixinghead[#MH].ReinigungskolbenGeregelt.GeneralParameters.Request := false;
           "PN_Mixinghead".Mixinghead[#MH].ReinigungskolbenGeregelt.Zeiten.Request := false;
           "PN_Mixinghead".Mixinghead[#MH].ReinigungskolbenGeregelt.Skalierung.Request := false;
           "PN_Mixinghead".Mixinghead[#MH].ReinigungskolbenGeregelt.Regelparameter.Request := false;
       END_IF;
       IF NOT "PN_Mixinghead".Mixinghead[#MH].ReinigungskolbenGesteuert.Active OR
           "PN_Mixinghead".Mixinghead[#MH].ReinigungskolbenGesteuert.Address = 0
       THEN
           "PN_Mixinghead".Mixinghead[#MH].ReinigungskolbenGesteuert.GeneralParameters.Request := false;
           "PN_Mixinghead".Mixinghead[#MH].ReinigungskolbenGesteuert.Zeiten.Request := false;
           "PN_Mixinghead".Mixinghead[#MH].ReinigungskolbenGesteuert.Skalierung.Request := false;
           "PN_Mixinghead".Mixinghead[#MH].ReinigungskolbenGesteuert.StufenAktivierung.Request := false;
           "PN_Mixinghead".Mixinghead[#MH].ReinigungskolbenGesteuert.StufenRückkehr.Request := false;
       END_IF;

       FOR #DB := 1 TO 8 DO
           IF NOT "PN_Mixinghead".Mixinghead[#MH].DüseBypass[#DB].Active THEN
               "PN_Mixinghead".Mixinghead[#MH].DüseBypass[#DB].Zeiten.Request := false;
           END_IF;
       END_FOR;

       // -----------------------------------
       // Mischkopf Analog   
       // -----------------------------------
       IF "PN_Mixinghead".Mixinghead[#MH].Analog.Active THEN
           #Address :=INT_TO_WORD("PN_Mixinghead".Mixinghead[#MH].Analog.Address);
           #ReturnValue := LOG2MOD(IOID := B#16#54, ADDR := #Address, HWID => #TempHWID);
           // Kommunikationsüberwachung
           // Nach einem Verbindungsabbruch werden die Telegramme automatisch verschickt.
           #Request := false;
           "CHCKPNCONN"(GOON := #GOON,
                        Active := "PN_Mixinghead".Mixinghead[#MH].Analog.Active,
                        Address := #TempHWID,
                        PN_Request := #Request,
                        PN_Fault := "PN_Mixinghead".Mixinghead[#MH].Analog.ChckConnFault,
                        DONE := "PN_Mixinghead".Mixinghead[#MH].Analog.ChckConnDone);

           IF #Request AND NOT "PN_Mixinghead".Mixinghead[#MH].Analog.ChckConnFault THEN
               "PN_Mixinghead".Mixinghead[#MH].Analog.Resourcen.Request := "PN_Mixinghead".Mixinghead[#MH].Analog.Active;
               "PN_Mixinghead".Mixinghead[#MH].Analog.Zeiten.Request := "PN_Mixinghead".Mixinghead[#MH].Analog.Active;
               "PN_Mixinghead".Mixinghead[#MH].Analog.Skalierung.Request := "PN_Mixinghead".Mixinghead[#MH].Analog.Active;
               "PN_Mixinghead".Mixinghead[#MH].Analog.StufenAktivierung.Request := "PN_Mixinghead".Mixinghead[#MH].Analog.Active;
               "PN_Mixinghead".Mixinghead[#MH].Analog.StufenRückkehr.Request := "PN_Mixinghead".Mixinghead[#MH].Analog.Active;
           END_IF;

           "WRREC_FC"(GOON := #GOON,
                      REQ := "PN_Mixinghead".Mixinghead[#MH].Analog.Resourcen.Request,
                      ACTIVE := "PN_Mixinghead".Mixinghead[#MH].Analog.Active,
                      ADDRESS := #TempHWID,
                      INDEX := #IDM_Mixinghead_Analog_Resourcen_Index,
                      LENGTH := #IDM_Mixinghead_Analog_Resourcen_Length,
                      WRREC_DONE => #t.DONE,
                      WRREC_BUSY => #t.BUSY,
                      WRREC_ERROR => #t.ERROR,
                      WRREC_STATUS => #t.STATUS,
                      RECORD := "PN_Mixinghead".Mixinghead[#MH].Analog.Resourcen.Data,
                      DONE := "PN_Mixinghead".Mixinghead[#MH].Analog.Resourcen.Transmitting);

           "WRREC_FC"(GOON := #GOON,
                      REQ := "PN_Mixinghead".Mixinghead[#MH].Analog.Zeiten.Request,
                      ACTIVE := "PN_Mixinghead".Mixinghead[#MH].Analog.Active,
                      ADDRESS := #TempHWID,
                      INDEX := #IDM_Mixinghead_Analog_Zeiten_Index,
                      LENGTH := #IDM_Mixinghead_Analog_Zeiten_Length,
                      WRREC_DONE => #t.DONE,
                      WRREC_BUSY => #t.BUSY,
                      WRREC_ERROR => #t.ERROR,
                      WRREC_STATUS => #t.STATUS,
                      RECORD := "PN_Mixinghead".Mixinghead[#MH].Analog.Zeiten.Data,
                      DONE := "PN_Mixinghead".Mixinghead[#MH].Analog.Zeiten.Transmitting);

           "WRREC_FC"(GOON := #GOON,
                      REQ := "PN_Mixinghead".Mixinghead[#MH].Analog.Skalierung.Request,
                      ACTIVE := "PN_Mixinghead".Mixinghead[#MH].Analog.Active,
                      ADDRESS := #TempHWID,
                      INDEX := #IDM_Mixinghead_Analog_Skalierung_Index,
                      LENGTH := #IDM_Mixinghead_Analog_Skalierung_Length,
                      WRREC_DONE => #t.DONE,
                      WRREC_BUSY => #t.BUSY,
                      WRREC_ERROR => #t.ERROR,
                      WRREC_STATUS => #t.STATUS,
                      RECORD := "PN_Mixinghead".Mixinghead[#MH].Analog.Skalierung.Data,
                      DONE := "PN_Mixinghead".Mixinghead[#MH].Analog.Skalierung.Transmitting);

           "WRREC_FC"(GOON := #GOON,
                      REQ := "PN_Mixinghead".Mixinghead[#MH].Analog.StufenAktivierung.Request,
                      ACTIVE := "PN_Mixinghead".Mixinghead[#MH].Analog.Active,
                      ADDRESS := #TempHWID,
                      INDEX := #IDM_Mixinghead_Analog_StufenAktivierung_Index,
                      LENGTH := #IDM_Mixinghead_Analog_StufenAktivierung_Length,
                      WRREC_DONE => #t.DONE,
                      WRREC_BUSY => #t.BUSY,
                      WRREC_ERROR => #t.ERROR,
                      WRREC_STATUS => #t.STATUS,
                      RECORD := "PN_Mixinghead".Mixinghead[#MH].Analog.StufenAktivierung.Data,
                      DONE := "PN_Mixinghead".Mixinghead[#MH].Analog.StufenAktivierung.Transmitting);

           "WRREC_FC"(GOON := #GOON,
                      REQ := "PN_Mixinghead".Mixinghead[#MH].Analog.StufenRückkehr.Request,
                      ACTIVE := "PN_Mixinghead".Mixinghead[#MH].Analog.Active,
                      ADDRESS := #TempHWID,
                      INDEX := #IDM_Mixinghead_Analog_StufenRückkehr_Index,
                      LENGTH := #IDM_Mixinghead_Analog_StufenRückkehr_Length,
                      WRREC_DONE => #t.DONE,
                      WRREC_BUSY => #t.BUSY,
                      WRREC_ERROR => #t.ERROR,
                      WRREC_STATUS => #t.STATUS,
                      RECORD := "PN_Mixinghead".Mixinghead[#MH].Analog.StufenRückkehr.Data,
                      DONE := "PN_Mixinghead".Mixinghead[#MH].Analog.StufenRückkehr.Transmitting);
       END_IF;

       // -----------------------------------
       // Mischkopf Digital   
       // -----------------------------------
       IF "PN_Mixinghead".Mixinghead[#MH].Digital.Active THEN
           #Address := INT_TO_WORD("PN_Mixinghead".Mixinghead[#MH].Digital.Address);
           #ReturnValue := LOG2MOD(IOID := B#16#54, ADDR := #Address, HWID => #TempHWID);
           // Kommunikationsüberwachung
           // Nach einem Verbindungsabbruch werden die Telegramme automatisch verschickt.
           #Request := false;
           "CHCKPNCONN"(
                        GOON := #GOON,
                        Active := "PN_Mixinghead".Mixinghead[#MH].Digital.Active,
                        Address := #TempHWID,
                        PN_Request := #Request,
                        PN_Fault := "PN_Mixinghead".Mixinghead[#MH].Digital.ChckConnFault,
                        DONE := "PN_Mixinghead".Mixinghead[#MH].Digital.ChckConnDone);

           IF #Request AND NOT "PN_Mixinghead".Mixinghead[#MH].Digital.ChckConnFault THEN
               "PN_Mixinghead".Mixinghead[#MH].Digital.GeneralParameters.Request := "PN_Mixinghead".Mixinghead[#MH].Digital.Active;
               "PN_Mixinghead".Mixinghead[#MH].Digital.Zeiten.Request := "PN_Mixinghead".Mixinghead[#MH].Digital.Active;
               "PN_Mixinghead".Mixinghead[#MH].Digital.Zeiten_2.Request := "PN_Mixinghead".Mixinghead[#MH].Digital.Active;
           END_IF;

           "WRREC_FC"(GOON := #GOON,
                      REQ := "PN_Mixinghead".Mixinghead[#MH].Digital.GeneralParameters.Request,
                      ADDRESS := #TempHWID,
                      INDEX := #IDM_Mixinghead_Digital_GeneralParameters_Index,
                      LENGTH := #IDM_Mixinghead_Digital_GeneralParameters_Length,
                      WRREC_DONE => #t.DONE,
                      WRREC_BUSY => #t.BUSY,
                      WRREC_ERROR => #t.ERROR,
                      WRREC_STATUS => #t.STATUS,
                      ACTIVE := "PN_Mixinghead".Mixinghead[#MH].Digital.Active,
                      RECORD := "PN_Mixinghead".Mixinghead[#MH].Digital.GeneralParameters.Data,
                      DONE := "PN_Mixinghead".Mixinghead[#MH].Digital.GeneralParameters.Transmitting);

           "WRREC_FC"(GOON := #GOON,
                      REQ := "PN_Mixinghead".Mixinghead[#MH].Digital.Zeiten.Request,
                      ADDRESS := #TempHWID,
                      INDEX := #IDM_Mixinghead_Digital_Zeiten_Index,
                      LENGTH := #IDM_Mixinghead_Digital_Zeiten_Length,
                      WRREC_DONE => #t.DONE,
                      WRREC_BUSY => #t.BUSY,
                      WRREC_ERROR => #t.ERROR,
                      WRREC_STATUS => #t.STATUS,
                      ACTIVE := "PN_Mixinghead".Mixinghead[#MH].Digital.Active,
                      RECORD := "PN_Mixinghead".Mixinghead[#MH].Digital.Zeiten.Data,
                      DONE := "PN_Mixinghead".Mixinghead[#MH].Digital.Zeiten.Transmitting);

           "WRREC_FC"(GOON := #GOON,
                      REQ := "PN_Mixinghead".Mixinghead[#MH].Digital.Zeiten_2.Request,
                      ADDRESS := #TempHWID,
                      INDEX := #IDM_Mixinghead_Digital_Zeiten_2_Index,
                      LENGTH := #IDM_Mixinghead_Digital_Zeiten_2_Length,
                      WRREC_DONE => #t.DONE,
                      WRREC_BUSY => #t.BUSY,
                      WRREC_ERROR => #t.ERROR,
                      WRREC_STATUS => #t.STATUS,
                      ACTIVE := "PN_Mixinghead".Mixinghead[#MH].Digital.Active,
                      RECORD := "PN_Mixinghead".Mixinghead[#MH].Digital.Zeiten_2.Data,
                      DONE := "PN_Mixinghead".Mixinghead[#MH].Digital.Zeiten_2.Transmitting);
       END_IF;

       // -----------------------------------
       // REINIGUNGSKOLBEN Digital   
       // -----------------------------------
       IF "PN_Mixinghead".Mixinghead[#MH].ReinigungskolbenDigital.Active THEN
           #Address := INT_TO_WORD("PN_Mixinghead".Mixinghead[#MH].ReinigungskolbenDigital.Address);
           #ReturnValue := LOG2MOD(IOID := B#16#54, ADDR := #Address, HWID => #TempHWID);
           // Kommunikationsüberwachung
           // Nach einem Verbindungsabbruch werden die Telegramme automatisch verschickt.
           #Request := false;
           "CHCKPNCONN"(GOON := #GOON,
                        Active := "PN_Mixinghead".Mixinghead[#MH].ReinigungskolbenDigital.Active,
                        Address := #TempHWID,
                        PN_Request := #Request,
                        PN_Fault := "PN_Mixinghead".Mixinghead[#MH].ReinigungskolbenDigital.ChckConnFault,
                        DONE := "PN_Mixinghead".Mixinghead[#MH].ReinigungskolbenDigital.ChckConnDone);

